FUNCTION_BLOCK "FB_Arg_Seq_1"   // FB2, GRAPH_PLUS
{ S7_Optimized_Access := 'TRUE' }
VERSION : 0.1
   VAR_INPUT
      OFF_SQ : Bool := false;   // Turn sequence off
      INIT_SQ : Bool := false;   // Set sequence to initial state
      ACK_EF : Bool := false;   // Acknowledge all errors and faults
      S_PREV : Bool := false;   // Output previous step in parameter S_NO
      S_NEXT : Bool := false;   // Indicate next step in parameter S_NO
      SW_AUTO : Bool := false;   // Automatic mode
      SW_TAP : Bool := false;   // Semiautomatic/switch with transition
      SW_TOP : Bool := false;   // Semiautomatic/ignore transition
      SW_MAN : Bool := false;   // Manual mode
      S_SEL : Int := 0;   // Select step to be output to S_NO
      S_ON : Bool := false;   // Activate step indicated in S_NO
      S_OFF : Bool := false;   // Deactivate step indicated S_NO
      T_PUSH : Bool := false;   // Enable transition to switch in semi automatic mode
      Start : Bool;
      stepTimes : Array[2..10] of Time;
      Model_Numb : Int := 3;
   END_VAR
   VAR_OUTPUT
      S_NO : Int := 0;   // Step number
      S_MORE : Bool := false;   // More steps are available and can be shown in S_NO
      S_ACTIVE : Bool := false;   // Step indicated in S_NO is active
      ERR_FLT : Bool := false;   // Interlock or supervision group error
      AUTO_ON : Bool := false;   // Automatic mode is active
      TAP_ON : Bool := false;   // Semiautomatic mode/step with transition enabled
      TOP_ON : Bool := false;   // Semiautomatic mode/ignore transition enabled
      MAN_ON : Bool := false;   // Manual mode is active
   END_VAR
   VAR
      HMI_INFO : Array[0..8] of UInt;
      IF_PAR : G7_IfParPlus_V6;
      RT_DATA : G7_RTDataPlus_V6;   // Internal data area
      Trans1 : G7_TransitionPlus_V6;   // Transition structure
      Trans2 : G7_TransitionPlus_V6;   // Transition structure
      Trans3 : G7_TransitionPlus_V6;   // Transition structure
      Trans4 : G7_TransitionPlus_V6;   // Transition structure
      Trans5 : G7_TransitionPlus_V6;   // Transition structure
      Trans6 : G7_TransitionPlus_V6;   // Transition structure
      Trans7 : G7_TransitionPlus_V6;   // Transition structure
      Trans8 : G7_TransitionPlus_V6;   // Transition structure
      Trans9 : G7_TransitionPlus_V6;   // Transition structure
      Trans10 : G7_TransitionPlus_V6;   // Transition structure
      Trans11 : G7_TransitionPlus_V6;   // Transition structure
      Trans12 : G7_TransitionPlus_V6;   // Transition structure
      Trans13 : G7_TransitionPlus_V6;   // Transition structure
      Trans14 : G7_TransitionPlus_V6;   // Transition structure
      Trans15 : G7_TransitionPlus_V6;   // Transition structure
      Trans16 : G7_TransitionPlus_V6;   // Transition structure
      Trans17 : G7_TransitionPlus_V6;   // Transition structure
      Trans18 : G7_TransitionPlus_V6;   // Transition structure
      Trans19 : G7_TransitionPlus_V6;   // Transition structure
      Trans21 : G7_TransitionPlus_V6;   // Transition structure
      "Step1: Init (Idle)" : G7_StepPlus_V6;   // Step structure
      Step2 : G7_StepPlus_V6;   // Step structure
      Step3 : G7_StepPlus_V6;   // Step structure
      Step4 : G7_StepPlus_V6;   // Step structure
      Step5 : G7_StepPlus_V6;   // Step structure
      Step6 : G7_StepPlus_V6;   // Step structure
      Step7 : G7_StepPlus_V6;   // Step structure
      Step8 : G7_StepPlus_V6;   // Step structure
      Step9 : G7_StepPlus_V6;   // Step structure
      Step10 : G7_StepPlus_V6;   // Step structure
      Step11 : G7_StepPlus_V6;   // Step structure
      Step12 : G7_StepPlus_V6;   // Step structure
      Step13 : G7_StepPlus_V6;   // Step structure
      Step14 : G7_StepPlus_V6;   // Step structure
      Step15 : G7_StepPlus_V6;   // Step structure
      Step16 : G7_StepPlus_V6;   // Step structure
      Step17 : G7_StepPlus_V6;   // Step structure
      Step18 : G7_StepPlus_V6;   // Step structure
      Step19 : G7_StepPlus_V6;   // Step structure
      SINI : Array[0..1] of USInt;
      LSTT : Array[0..19] of USInt;
      ATAJ : Array[0..19] of USInt;
      ATAB : Array[0..19] of USInt;
      PSTT : Array[0..19] of USInt;
      NSTT : Array[0..19] of USInt;
      ASSJ : Array[0..18] of USInt;
      ASSB : Array[0..18] of USInt;
      PTTS : Array[0..18] of USInt;
      NTTS : Array[0..18] of USInt;
      SW_SQTS : Array[0..18] of USInt;
      SWITCH : Array[0..1] of USInt;
      TVX : Array[0..3] of USInt;
      TTX : Array[0..3] of USInt;
      TSX : Array[0..1] of USInt;
      S00X : Array[0..1] of USInt;
      SOFFX : Array[0..1] of USInt;
      SONX : Array[0..1] of USInt;
      SAX : Array[0..1] of USInt;
      SERRX : Array[0..19] of USInt;
      SMX : Array[0..19] of USInt;
      S0X : Array[0..19] of USInt;
      S1X : Array[0..19] of USInt;
      IL_ALARM_INST : Diag_Alarm;
      SUP_ALARM_INST : Diag_Alarm;
      STEP_TIME_ALARM_INST : Diag_Alarm;
      IEC_TIMER_INST : IEC_TIMER;
      TRANSACTION_FLAG : Bool := false;
   END_VAR
   // SINI[0] := 2;
   // LSTT[0] := 255;
   // LSTT[1] := 255;
   // LSTT[2] := 255;
   // ATAJ[1] := 1;
   // ATAJ[2] := 2;
   // ATAJ[3] := 3;
   // ATAB[1] := 1;
   // ATAB[2] := 2;
   // ATAB[3] := 3;
   // PSTT[1] := 1;
   // PSTT[2] := 2;
   // PSTT[3] := 3;
   // NSTT[0] := 1;
   // NSTT[1] := 2;
   // NSTT[2] := 3;
   // ASSJ[1] := 1;
   // ASSJ[2] := 2;
   // ASSJ[3] := 3;
   // ASSB[1] := 1;
   // ASSB[2] := 2;
   // ASSB[3] := 3;
   // PTTS[0] := 255;
   // PTTS[2] := 1;
   // PTTS[3] := 2;
   // NTTS[1] := 1;
   // NTTS[2] := 2;
   // NTTS[3] := 3;
   // TVX[0] := 16#1;
   // TTX[0] := 16#1;
   // TSX[0] := 16#1;
   // S00X[0] := 16#1;
   // SOFFX[0] := 16#1;
   // SONX[0] := 16#1;
   // SAX[0] := 16#1;
   // SERRX[0] := 16#1;
   // SMX[0] := 16#1;
   // S0X[0] := 16#1;
   // S1X[0] := 16#1;
   // LSTT[3] := 255;
   // LSTT[4] := 255;
   // LSTT[5] := 255;
   // LSTT[6] := 255;
   // LSTT[7] := 255;
   // LSTT[8] := 255;
   // ATAJ[4] := 4;
   // ATAJ[5] := 5;
   // ATAJ[6] := 6;
   // ATAJ[7] := 7;
   // ATAJ[8] := 8;
   // ATAJ[9] := 9;
   // ATAB[4] := 4;
   // ATAB[5] := 5;
   // ATAB[6] := 6;
   // ATAB[7] := 7;
   // ATAB[8] := 8;
   // ATAB[9] := 9;
   // PSTT[4] := 4;
   // PSTT[5] := 5;
   // PSTT[6] := 6;
   // PSTT[7] := 7;
   // PSTT[8] := 8;
   // PSTT[9] := 9;
   // NSTT[3] := 4;
   // NSTT[4] := 5;
   // NSTT[5] := 6;
   // NSTT[6] := 7;
   // NSTT[7] := 8;
   // NSTT[8] := 9;
   // ASSJ[4] := 4;
   // ASSJ[5] := 5;
   // ASSJ[6] := 6;
   // ASSJ[7] := 7;
   // ASSJ[8] := 8;
   // ASSJ[9] := 9;
   // ASSB[4] := 4;
   // ASSB[5] := 5;
   // ASSB[6] := 6;
   // ASSB[7] := 7;
   // ASSB[8] := 8;
   // ASSB[9] := 9;
   // PTTS[4] := 3;
   // PTTS[5] := 4;
   // PTTS[6] := 5;
   // PTTS[7] := 6;
   // PTTS[8] := 7;
   // PTTS[9] := 8;
   // NTTS[4] := 4;
   // NTTS[5] := 5;
   // NTTS[6] := 6;
   // NTTS[7] := 7;
   // NTTS[8] := 8;
   // NTTS[9] := 9;
   // LSTT[10] := 255;
   // LSTT[11] := 255;
   // LSTT[12] := 255;
   // LSTT[13] := 255;
   // LSTT[14] := 255;
   // LSTT[15] := 255;
   // LSTT[16] := 255;
   // LSTT[17] := 255;
   // LSTT[18] := 255;
   // ATAJ[10] := 10;
   // ATAJ[11] := 11;
   // ATAJ[12] := 12;
   // ATAJ[13] := 13;
   // ATAJ[14] := 14;
   // ATAJ[15] := 15;
   // ATAJ[16] := 16;
   // ATAJ[17] := 17;
   // ATAJ[18] := 18;
   // ATAJ[19] := 19;
   // ATAB[0] := 10;
   // ATAB[11] := 11;
   // ATAB[12] := 12;
   // ATAB[13] := 13;
   // ATAB[14] := 14;
   // ATAB[15] := 15;
   // ATAB[16] := 16;
   // ATAB[17] := 17;
   // ATAB[18] := 18;
   // ATAB[19] := 19;
   // PSTT[11] := 10;
   // PSTT[12] := 11;
   // PSTT[13] := 12;
   // PSTT[14] := 13;
   // PSTT[15] := 14;
   // PSTT[16] := 15;
   // PSTT[17] := 16;
   // PSTT[18] := 17;
   // PSTT[19] := 18;
   // NSTT[10] := 10;
   // NSTT[11] := 11;
   // NSTT[12] := 12;
   // NSTT[13] := 13;
   // NSTT[14] := 14;
   // NSTT[15] := 15;
   // NSTT[16] := 16;
   // NSTT[17] := 17;
   // NSTT[18] := 18;
   // ASSJ[10] := 10;
   // ASSJ[11] := 11;
   // ASSJ[12] := 12;
   // ASSJ[13] := 13;
   // ASSJ[14] := 14;
   // ASSJ[15] := 15;
   // ASSJ[16] := 16;
   // ASSJ[17] := 17;
   // ASSJ[18] := 18;
   // ASSB[10] := 10;
   // ASSB[11] := 11;
   // ASSB[12] := 12;
   // ASSB[13] := 13;
   // ASSB[14] := 14;
   // ASSB[15] := 15;
   // ASSB[16] := 16;
   // ASSB[17] := 17;
   // ASSB[18] := 18;
   // PTTS[10] := 10;
   // PTTS[11] := 11;
   // PTTS[12] := 12;
   // PTTS[13] := 13;
   // PTTS[14] := 14;
   // PTTS[15] := 15;
   // PTTS[16] := 16;
   // PTTS[17] := 17;
   // PTTS[18] := 18;
   // NTTS[10] := 11;
   // NTTS[11] := 12;
   // NTTS[12] := 13;
   // NTTS[13] := 14;
   // NTTS[14] := 15;
   // NTTS[15] := 16;
   // NTTS[16] := 17;
   // NTTS[17] := 18;
   // NTTS[18] := 19;
   // SW_SQTS[1] := 1;
   // SW_SQTS[2] := 1;
   // SW_SQTS[3] := 1;
   // SW_SQTS[4] := 1;
   // SW_SQTS[5] := 1;
   // SW_SQTS[6] := 1;
   // SW_SQTS[7] := 1;
   // SW_SQTS[8] := 1;
   // SW_SQTS[9] := 1;
   // SW_SQTS[10] := 2;
   // SW_SQTS[11] := 2;
   // SW_SQTS[12] := 2;
   // SW_SQTS[13] := 2;
   // SW_SQTS[14] := 2;
   // SW_SQTS[15] := 2;
   // SW_SQTS[16] := 2;
   // SW_SQTS[17] := 2;
   // SW_SQTS[18] := 2;
BEGIN
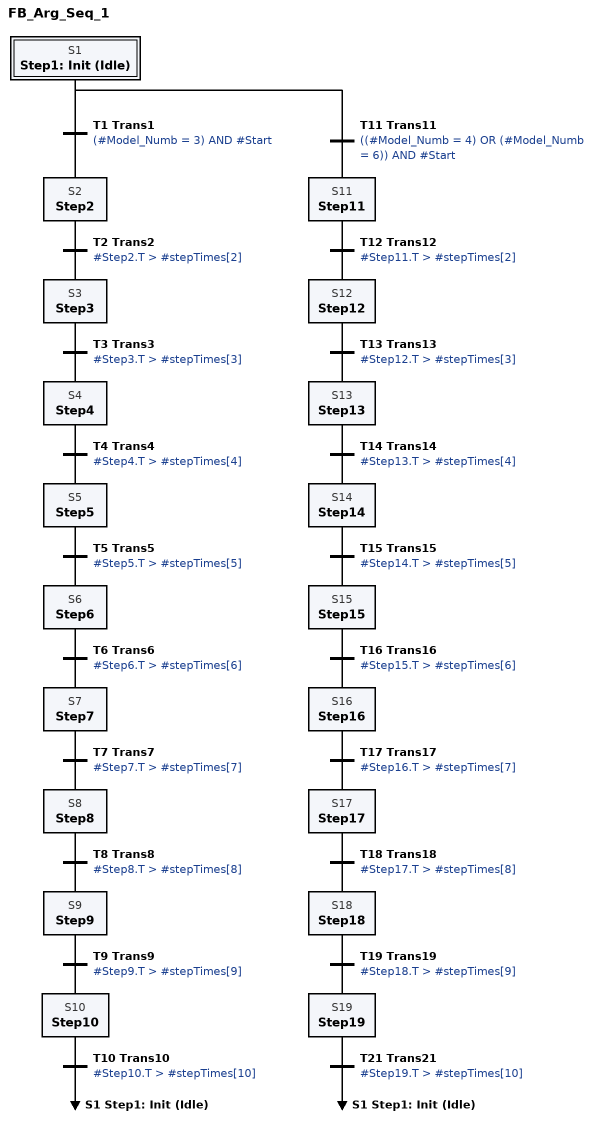
   // sequencer 1
   INITIAL_STEP "Step1: Init (Idle)":   // S1, max time T#10S, warning time T#7S
   END_STEP
   TRANSITION Trans1 FROM "Step1: Init (Idle)" TO Step2   // T1
      := (#Model_Numb = 3) AND #Start;
   END_TRANSITION
   TRANSITION Trans11 FROM "Step1: Init (Idle)" TO Step11   // T11
      := ((#Model_Numb = 4) OR (#Model_Numb = 6)) AND #Start;
   END_TRANSITION
   STEP Step2:   // S2, max time T#10S, warning time T#7S
   END_STEP
   TRANSITION Trans2 FROM Step2 TO Step3   // T2
      := #Step2.T > #stepTimes[2];
   END_TRANSITION
   STEP Step3:   // S3, max time T#10S, warning time T#7S
   END_STEP
   TRANSITION Trans3 FROM Step3 TO Step4   // T3
      := #Step3.T > #stepTimes[3];
   END_TRANSITION
   STEP Step4:   // S4, max time T#10S, warning time T#7S
   END_STEP
   TRANSITION Trans4 FROM Step4 TO Step5   // T4
      := #Step4.T > #stepTimes[4];
   END_TRANSITION
   STEP Step5:   // S5, max time T#10S, warning time T#7S
   END_STEP
   TRANSITION Trans5 FROM Step5 TO Step6   // T5
      := #Step5.T > #stepTimes[5];
   END_TRANSITION
   STEP Step6:   // S6, max time T#10S, warning time T#7S
   END_STEP
   TRANSITION Trans6 FROM Step6 TO Step7   // T6
      := #Step6.T > #stepTimes[6];
   END_TRANSITION
   STEP Step7:   // S7, max time T#10S, warning time T#7S
   END_STEP
   TRANSITION Trans7 FROM Step7 TO Step8   // T7
      := #Step7.T > #stepTimes[7];
   END_TRANSITION
   STEP Step8:   // S8, max time T#10S, warning time T#7S
   END_STEP
   TRANSITION Trans8 FROM Step8 TO Step9   // T8
      := #Step8.T > #stepTimes[8];
   END_TRANSITION
   STEP Step9:   // S9, max time T#10S, warning time T#7S
   END_STEP
   TRANSITION Trans9 FROM Step9 TO Step10   // T9
      := #Step9.T > #stepTimes[9];
   END_TRANSITION
   STEP Step10:   // S10, max time T#10S, warning time T#7S
   END_STEP
   TRANSITION Trans10 FROM Step10 TO "Step1: Init (Idle)"   // T10, jump
      := #Step10.T > #stepTimes[10];
   END_TRANSITION
   STEP Step11:   // S11, max time T#10S, warning time T#7S
   END_STEP
   TRANSITION Trans12 FROM Step11 TO Step12   // T12
      := #Step11.T > #stepTimes[2];
   END_TRANSITION
   STEP Step12:   // S12, max time T#10S, warning time T#7S
   END_STEP
   TRANSITION Trans13 FROM Step12 TO Step13   // T13
      := #Step12.T > #stepTimes[3];
   END_TRANSITION
   STEP Step13:   // S13, max time T#10S, warning time T#7S
   END_STEP
   TRANSITION Trans14 FROM Step13 TO Step14   // T14
      := #Step13.T > #stepTimes[4];
   END_TRANSITION
   STEP Step14:   // S14, max time T#10S, warning time T#7S
   END_STEP
   TRANSITION Trans15 FROM Step14 TO Step15   // T15
      := #Step14.T > #stepTimes[5];
   END_TRANSITION
   STEP Step15:   // S15, max time T#10S, warning time T#7S
   END_STEP
   TRANSITION Trans16 FROM Step15 TO Step16   // T16
      := #Step15.T > #stepTimes[6];
   END_TRANSITION
   STEP Step16:   // S16, max time T#10S, warning time T#7S
   END_STEP
   TRANSITION Trans17 FROM Step16 TO Step17   // T17
      := #Step16.T > #stepTimes[7];
   END_TRANSITION
   STEP Step17:   // S17, max time T#10S, warning time T#7S
   END_STEP
   TRANSITION Trans18 FROM Step17 TO Step18   // T18
      := #Step17.T > #stepTimes[8];
   END_TRANSITION
   STEP Step18:   // S18, max time T#10S, warning time T#7S
   END_STEP
   TRANSITION Trans19 FROM Step18 TO Step19   // T19
      := #Step18.T > #stepTimes[9];
   END_TRANSITION
   STEP Step19:   // S19, max time T#10S, warning time T#7S
   END_STEP
   TRANSITION Trans21 FROM Step19 TO "Step1: Init (Idle)"   // T21, jump
      := #Step19.T > #stepTimes[10];
   END_TRANSITION
END_FUNCTION_BLOCK

FUNCTION "FC_ARG_1" : Void   // FC1, FBD
{ S7_Optimized_Access := 'TRUE' }
VERSION : 0.1
   VAR_OUTPUT
      Ready_new_car : Bool;
   END_VAR
   VAR_TEMP
      stepTimes : Array[2..10] of Time;
      i : Int;
      Random_Time : Time;   // Random Time between 0sec to 10sec
      Start : Bool;
      Stop : Bool;
      status1_RandFunc : Word;
      status2_RandFunc : Word;
      temp : Byte;
      error_RandFunc : Bool;
   END_VAR
   VAR CONSTANT
      sequenceNO : Int := 9;
   END_VAR
BEGIN

REGION Network 1 (SCL): Man Mode Data Handling
   IF "DB_Process_Var".Man_Mode = TRUE THEN
       "DB_Process_Var".Car_Type_Selected := "DB_HMI".dropdown_selection;
   END_IF;
END_REGION

REGION Network 2 (SCL): Auto Mode Data Handling
   IF "DB_Process_Var".Auto_Mode = TRUE THEN
       "DB_HMI".dropdown_selection := 0;
       "DB_Process_Var".Car_Type_Selected := "DB_PLC5_Receiving".ReceivingBoxForward.Type;
   END_IF;
   IF "DB_HMI".ARG1_Seq1_Cmd_Auto OR "DB_HMI".Global_Cmd_Auto THEN
       "DB_HMI".dropdown_selection := 0;
       "DB_Process_Var".Car_Type_Selected := 0;
   END_IF;
END_REGION

REGION Network 3 (SCL): Load Time Date based on Car Type
       CASE "DB_Process_Var".Car_Type_Selected OF
           3:
               "DB_Profile"."time" := "DB_Profile".time_Red;
           4:
               "DB_Profile"."time" := "DB_Profile".time_Green;
           6:
               "DB_Profile"."time" := "DB_Profile".time_Blue;
       END_CASE;
END_REGION

REGION Network 4 (SCL): Switch from selected to inProduction
   IF "IDB_Arg_Seq_1_DB".Trans1.TS = TRUE OR "IDB_Arg_Seq_1_DB".Trans11.TS = TRUE THEN
       IF "DB_Process_Var".Car_Type_Selected = 3 THEN
           "DB_Process_Var".Car_Type_inProduction := 3;
           "DB_Process_Var".Car_Type_inProduction_Text := 'Red';
           "DB_HMI".ARG1_Seq1_inProduction := 3;
       ELSIF "DB_Process_Var".Car_Type_Selected = 4 THEN
           "DB_Process_Var".Car_Type_inProduction := 4;
           "DB_Process_Var".Car_Type_inProduction_Text := 'Green';
           "DB_HMI".ARG1_Seq1_inProduction := 4;
       ELSIF "DB_Process_Var".Car_Type_Selected = 6 THEN
           "DB_Process_Var".Car_Type_inProduction := 6;
           "DB_Process_Var".Car_Type_inProduction_Text := 'Blue';
           "DB_HMI".ARG1_Seq1_inProduction := 6;
       END_IF;
   END_IF;
END_REGION

REGION Network 5 (SCL): Create Random Time Values for the selected Steps
   IF "IDB_Arg_Seq_1_DB".Trans1.TS = TRUE OR "IDB_Arg_Seq_1_DB".Trans11.TS = TRUE THEN
       FOR #i := 2 TO 10 DO
           //Red
           IF "DB_HMI".ARG1_Seq1_DelaySelect_Red[#i] = TRUE THEN;
               "DB_Sim".Delta_T_Red[#i] := "LGF_RandomRange_Dint"(minValue := 0, maxValue := 10000, error => #error_RandFunc, status => #status1_RandFunc, subfunctionStatus => #status2_RandFunc);
           ELSE
               "DB_Sim".Delta_T_Red[#i] := T#0s;
           END_IF;
           //Green
           IF "DB_HMI".ARG1_Seq1_DelaySelect_Green[#i] = TRUE THEN
               "DB_Sim".Delta_T_Green[#i] := "LGF_RandomRange_Dint"(minValue := 0, maxValue := 10000, error => #error_RandFunc, status => #status1_RandFunc, subfunctionStatus => #status2_RandFunc);
           ELSE
               "DB_Sim".Delta_T_Green[#i] := T#0s;
           END_IF;
           //Blue
           IF "DB_HMI".ARG1_Seq1_DelaySelect_Blue[#i] = TRUE THEN
               "DB_Sim".Delta_T_Blue[#i] := "LGF_RandomRange_Dint"(minValue := 0, maxValue := 10000, error => #error_RandFunc, status => #status1_RandFunc, subfunctionStatus => #status2_RandFunc);
           ELSE
               "DB_Sim".Delta_T_Blue[#i] := T#0s;
           END_IF;
       END_FOR;
   END_IF;

   IF "DB_HMI".ARG1_Seq1_Cmd_DelayReset = TRUE THEN
       FOR #i := 2 TO 10 DO
           "DB_HMI".ARG1_Seq1_DelaySelect_Red[#i] := false;
           "DB_HMI".ARG1_Seq1_DelaySelect_Green[#i] := false;
           "DB_HMI".ARG1_Seq1_DelaySelect_Blue[#i] := false;
       END_FOR;
   END_IF;
END_REGION

REGION Network 6 (SCL): Add Delay Time to Step Time
   FOR #i := 2 TO 10 DO
       IF "DB_HMI".dropdown_selection = 3 OR "DB_PLC5_Receiving".ReceivingBoxForward.Type = 3 THEN
           "DB_Process_Var".Step_Times[#i] := T_ADD(IN1 := "DB_Profile"."time"[#i], IN2 := "DB_Sim".Delta_T_Red[#i]);
       ELSIF "DB_HMI".dropdown_selection = 4 OR "DB_PLC5_Receiving".ReceivingBoxForward.Type = 4 THEN
           "DB_Process_Var".Step_Times[#i] := T_ADD(IN1 := "DB_Profile"."time"[#i], IN2 := "DB_Sim".Delta_T_Green[#i]);
       ELSIF "DB_HMI".dropdown_selection = 6 OR "DB_PLC5_Receiving".ReceivingBoxForward.Type = 6 THEN
           "DB_Process_Var".Step_Times[#i] := T_ADD(IN1 := "DB_Profile"."time"[#i], IN2 := "DB_Sim".Delta_T_Blue[#i]);
       END_IF;
   END_FOR;
END_REGION

REGION Network 7: Auto Mode select
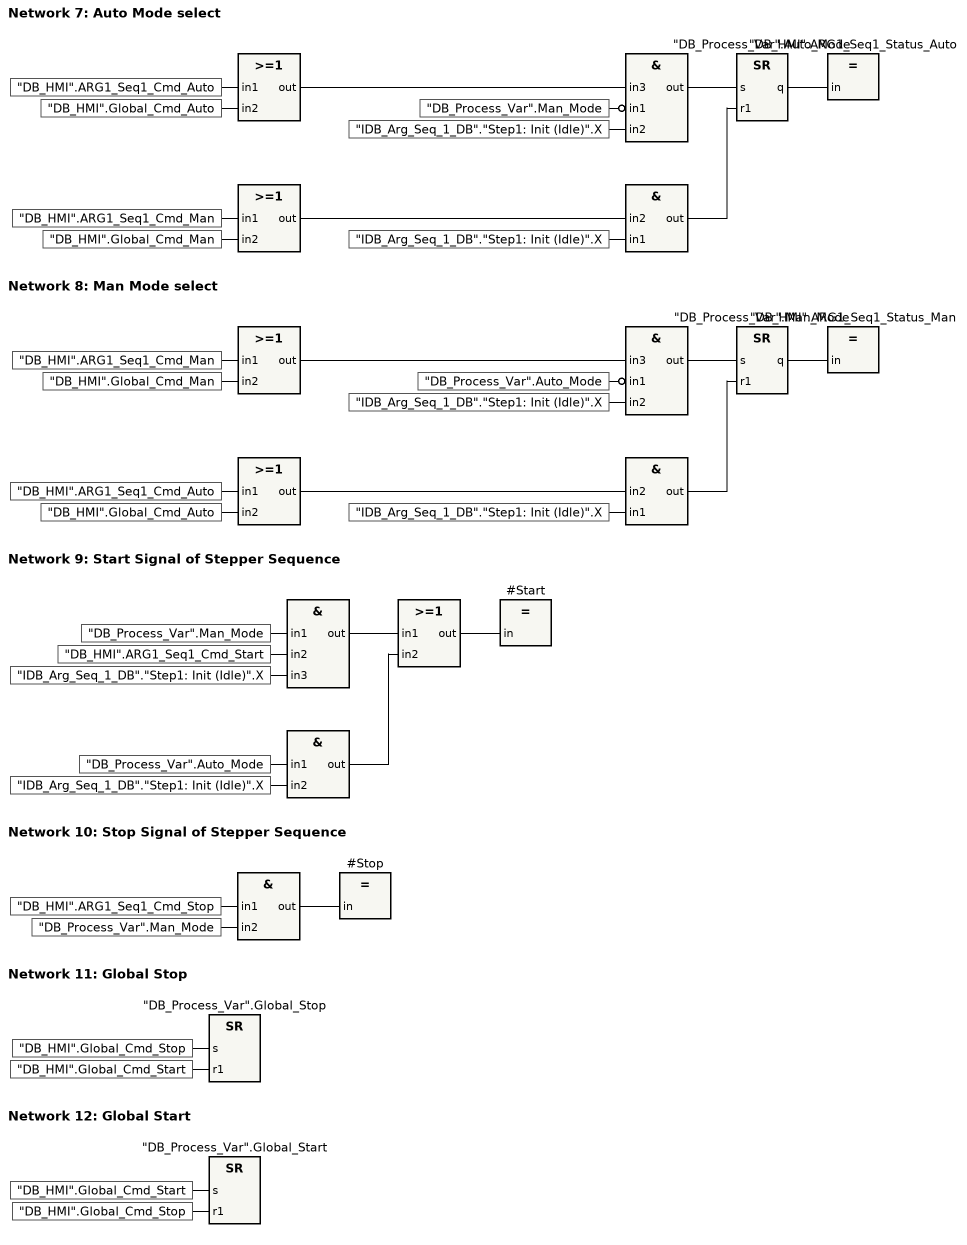
   IF ("DB_HMI".ARG1_Seq1_Cmd_Auto OR "DB_HMI".Global_Cmd_Auto) AND NOT "DB_Process_Var".Man_Mode AND "IDB_Arg_Seq_1_DB"."Step1: Init (Idle)".X THEN
       "DB_Process_Var".Auto_Mode := TRUE;   // SR flip-flop
   END_IF;
   IF ("DB_HMI".ARG1_Seq1_Cmd_Man OR "DB_HMI".Global_Cmd_Man) AND "IDB_Arg_Seq_1_DB"."Step1: Init (Idle)".X THEN
       "DB_Process_Var".Auto_Mode := FALSE;
   END_IF;
   "DB_HMI".ARG1_Seq1_Status_Auto := "DB_Process_Var".Auto_Mode;
END_REGION

REGION Network 8: Man Mode select
   IF ("DB_HMI".ARG1_Seq1_Cmd_Man OR "DB_HMI".Global_Cmd_Man) AND NOT "DB_Process_Var".Auto_Mode AND "IDB_Arg_Seq_1_DB"."Step1: Init (Idle)".X THEN
       "DB_Process_Var".Man_Mode := TRUE;   // SR flip-flop
   END_IF;
   IF ("DB_HMI".ARG1_Seq1_Cmd_Auto OR "DB_HMI".Global_Cmd_Auto) AND "IDB_Arg_Seq_1_DB"."Step1: Init (Idle)".X THEN
       "DB_Process_Var".Man_Mode := FALSE;
   END_IF;
   "DB_HMI".ARG1_Seq1_Status_Man := "DB_Process_Var".Man_Mode;
END_REGION

REGION Network 9: Start Signal of Stepper Sequence
   #Start := ("DB_Process_Var".Man_Mode AND "DB_HMI".ARG1_Seq1_Cmd_Start AND "IDB_Arg_Seq_1_DB"."Step1: Init (Idle)".X) OR ("DB_Process_Var".Auto_Mode AND "IDB_Arg_Seq_1_DB"."Step1: Init (Idle)".X);
END_REGION

REGION Network 10: Stop Signal of Stepper Sequence
   #Stop := "DB_HMI".ARG1_Seq1_Cmd_Stop AND "DB_Process_Var".Man_Mode;
END_REGION

REGION Network 11: Global Stop
   IF "DB_HMI".Global_Cmd_Stop THEN
       "DB_Process_Var".Global_Stop := TRUE;   // SR flip-flop
   END_IF;
   IF "DB_HMI".Global_Cmd_Start THEN "DB_Process_Var".Global_Stop := FALSE; END_IF;
END_REGION

REGION Network 12: Global Start
   IF "DB_HMI".Global_Cmd_Start THEN
       "DB_Process_Var".Global_Start := TRUE;   // SR flip-flop
   END_IF;
   IF "DB_HMI".Global_Cmd_Stop THEN "DB_Process_Var".Global_Start := FALSE; END_IF;
END_REGION

REGION Network 13 (SCL): Reset Type Selection
   IF "DB_HMI".ARG1_Seq1_Cmd_Stop = TRUE THEN
       "DB_PLC5_Receiving".ReceivingBoxForward.Type := 0;
       "DB_HMI".ARG1_Seq1_inProduction := 0;
       "DB_Process_Var".ReadyNewCar := TRUE;
   END_IF;
END_REGION

REGION Network 14: Call FB with Stepper Sequence
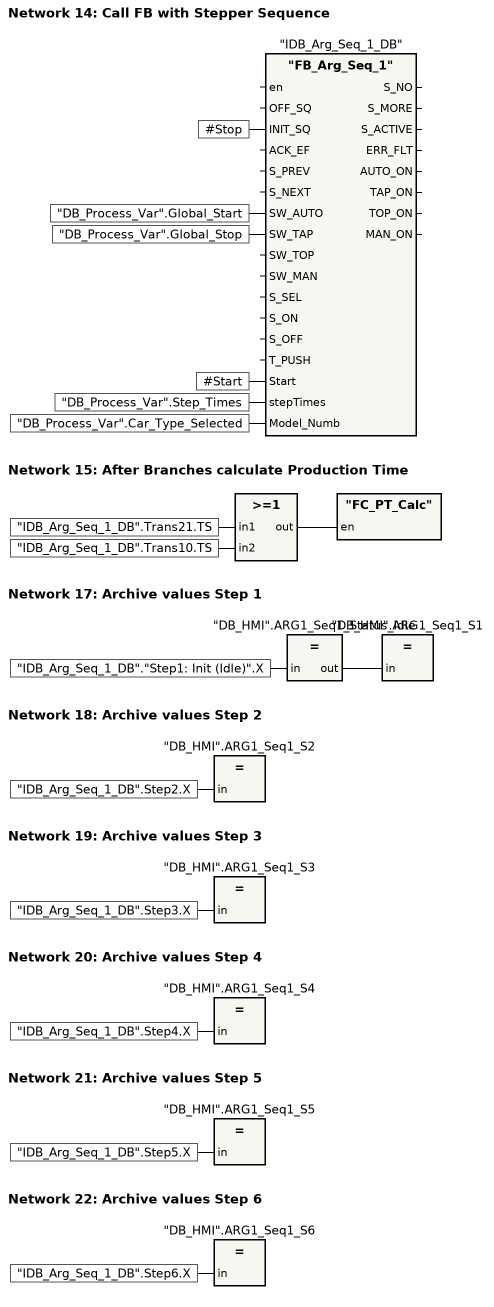
   "IDB_Arg_Seq_1_DB"(INIT_SQ := #Stop,   // "FB_Arg_Seq_1"
                      SW_AUTO := "DB_Process_Var".Global_Start,
                      SW_TAP := "DB_Process_Var".Global_Stop,
                      Start := #Start,
                      stepTimes := "DB_Process_Var".Step_Times,
                      Model_Numb := "DB_Process_Var".Car_Type_Selected);
END_REGION

REGION Network 15: After Branches calculate Production Time
   IF "IDB_Arg_Seq_1_DB".Trans21.TS OR "IDB_Arg_Seq_1_DB".Trans10.TS THEN "FC_PT_Calc"(); END_IF;
END_REGION

REGION Network 16 (SCL): Send Idle to previous Station
   IF "IDB_Arg_Seq_1_DB"."Step1: Init (Idle)".X = TRUE THEN
       "DB_PLC5_Sending".SendBox.Station_Idle := TRUE;
   ELSE
       "DB_PLC5_Sending".SendBox.Station_Idle := FALSE;
   END_IF;
END_REGION

REGION Network 17: Archive values Step 1
   "DB_HMI".ARG1_Seq1_Status_Idle := "IDB_Arg_Seq_1_DB"."Step1: Init (Idle)".X;
   "DB_HMI".ARG1_Seq1_S1 := "IDB_Arg_Seq_1_DB"."Step1: Init (Idle)".X;
END_REGION

REGION Network 18: Archive values Step 2
   "DB_HMI".ARG1_Seq1_S2 := "IDB_Arg_Seq_1_DB".Step2.X;
END_REGION

REGION Network 19: Archive values Step 3
   "DB_HMI".ARG1_Seq1_S3 := "IDB_Arg_Seq_1_DB".Step3.X;
END_REGION

REGION Network 20: Archive values Step 4
   "DB_HMI".ARG1_Seq1_S4 := "IDB_Arg_Seq_1_DB".Step4.X;
END_REGION

REGION Network 21: Archive values Step 5
   "DB_HMI".ARG1_Seq1_S5 := "IDB_Arg_Seq_1_DB".Step5.X;
END_REGION

REGION Network 22: Archive values Step 6
   "DB_HMI".ARG1_Seq1_S6 := "IDB_Arg_Seq_1_DB".Step6.X;
END_REGION

REGION Network 23: Archive values Step 7
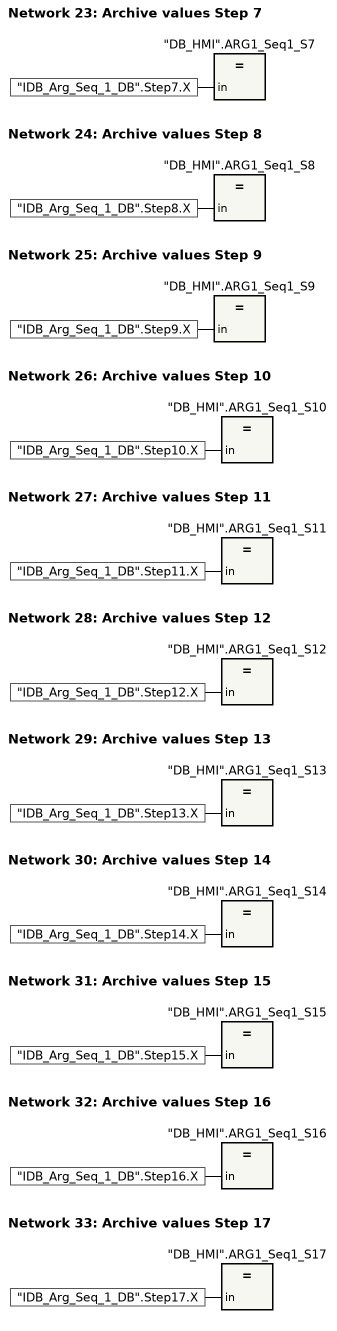
   "DB_HMI".ARG1_Seq1_S7 := "IDB_Arg_Seq_1_DB".Step7.X;
END_REGION

REGION Network 24: Archive values Step 8
   "DB_HMI".ARG1_Seq1_S8 := "IDB_Arg_Seq_1_DB".Step8.X;
END_REGION

REGION Network 25: Archive values Step 9
   "DB_HMI".ARG1_Seq1_S9 := "IDB_Arg_Seq_1_DB".Step9.X;
END_REGION

REGION Network 26: Archive values Step 10
   "DB_HMI".ARG1_Seq1_S10 := "IDB_Arg_Seq_1_DB".Step10.X;
END_REGION

REGION Network 27: Archive values Step 11
   "DB_HMI".ARG1_Seq1_S11 := "IDB_Arg_Seq_1_DB".Step11.X;
END_REGION

REGION Network 28: Archive values Step 12
   "DB_HMI".ARG1_Seq1_S12 := "IDB_Arg_Seq_1_DB".Step12.X;
END_REGION

REGION Network 29: Archive values Step 13
   "DB_HMI".ARG1_Seq1_S13 := "IDB_Arg_Seq_1_DB".Step13.X;
END_REGION

REGION Network 30: Archive values Step 14
   "DB_HMI".ARG1_Seq1_S14 := "IDB_Arg_Seq_1_DB".Step14.X;
END_REGION

REGION Network 31: Archive values Step 15
   "DB_HMI".ARG1_Seq1_S15 := "IDB_Arg_Seq_1_DB".Step15.X;
END_REGION

REGION Network 32: Archive values Step 16
   "DB_HMI".ARG1_Seq1_S16 := "IDB_Arg_Seq_1_DB".Step16.X;
END_REGION

REGION Network 33: Archive values Step 17
   "DB_HMI".ARG1_Seq1_S17 := "IDB_Arg_Seq_1_DB".Step17.X;
END_REGION

REGION Network 34: Archive values Step 18
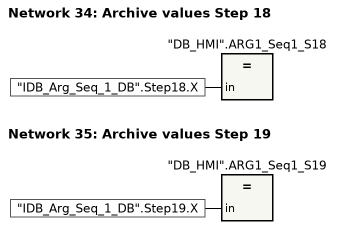
   "DB_HMI".ARG1_Seq1_S18 := "IDB_Arg_Seq_1_DB".Step18.X;
END_REGION

REGION Network 35: Archive values Step 19
   "DB_HMI".ARG1_Seq1_S19 := "IDB_Arg_Seq_1_DB".Step19.X;
END_REGION

REGION Network 36 (SCL): Set Busy
   IF
       "IDB_Arg_Seq_1_DB".Step2.X OR
       "IDB_Arg_Seq_1_DB".Step3.X OR
       "IDB_Arg_Seq_1_DB".Step4.X OR
       "IDB_Arg_Seq_1_DB".Step5.X OR
       "IDB_Arg_Seq_1_DB".Step6.X OR
       "IDB_Arg_Seq_1_DB".Step7.X OR
       "IDB_Arg_Seq_1_DB".Step8.X OR
       "IDB_Arg_Seq_1_DB".Step9.X OR
       "IDB_Arg_Seq_1_DB".Step10.X OR
       "IDB_Arg_Seq_1_DB".Step11.X OR
       "IDB_Arg_Seq_1_DB".Step12.X OR
       "IDB_Arg_Seq_1_DB".Step13.X OR
       "IDB_Arg_Seq_1_DB".Step14.X OR
       "IDB_Arg_Seq_1_DB".Step15.X OR
       "IDB_Arg_Seq_1_DB".Step16.X OR
       "IDB_Arg_Seq_1_DB".Step17.X OR
       "IDB_Arg_Seq_1_DB".Step18.X OR
       "IDB_Arg_Seq_1_DB".Step19.X THEN
       "DB_HMI".ARG1_Seq1_Status_Busy := TRUE;
   ELSIF "IDB_Arg_Seq_1_DB"."Step1: Init (Idle)".X THEN
       "DB_HMI".ARG1_Seq1_Status_Busy := FALSE;
   END_IF;
END_REGION

REGION Network 37 (SCL): When Stepper Sequence runs completely
   IF "IDB_Arg_Seq_1_DB".Trans10.TS = TRUE OR "IDB_Arg_Seq_1_DB".Trans21.TS = TRUE THEN
       "DB_Process_Var".Branch_Complete := TRUE;
       "DB_Process_Var".Car_Type_Ready := "DB_Process_Var".Car_Type_inProduction;
       "DB_Process_Var".Car_Type_inProduction := 0;
       "DB_Process_Var".Car_Type_inProduction_Text := '';
       "DB_Process_Var".Car_ReadyToShift := TRUE;
       "DB_HMI".ARG1_Seq1_inProduction := 0;
   END_IF;
   IF "IDB_Arg_Seq_1_DB".Trans1.TS = TRUE OR "IDB_Arg_Seq_1_DB".Trans11.TS = TRUE THEN
       "DB_Process_Var".Branch_Complete := FALSE;
       "DB_Process_Var".ReadyNewCar := 0;
   END_IF;
END_REGION

REGION Network 38 (SCL): Write Data in the Sending Box
   //IF "DB_Process_Var".Branch_Complete = TRUE AND "DB_PLC5_Receiving".ReceivingBox.Station_Idle = TRUE THEN
   IF "IDB_Arg_Seq_1_DB".Trans10.TS = TRUE OR "IDB_Arg_Seq_1_DB".Trans21.TS = TRUE THEN
       "DB_PLC5_Sending".SendBoxForward.Planned_PT_Red := "DB_HMI".ARG1_Seq1_Calculated_PT_Red;
       "DB_PLC5_Sending".SendBoxForward.Planned_PT_Green := "DB_HMI".ARG1_Seq1_Calculated_PT_Green;
       "DB_PLC5_Sending".SendBoxForward.Planned_PT_Blue := "DB_HMI".ARG1_Seq1_Calculated_PT_Blue;

       "DB_PLC5_Sending".SendBoxForward.Measuered_PT_Red := "DB_HMI".ARG1_Seq1_Messured_PT_Red;
       "DB_PLC5_Sending".SendBoxForward.Measuered_PT_Green := "DB_HMI".ARG1_Seq1_Messured_PT_Green;
       "DB_PLC5_Sending".SendBoxForward.Measuered_PT_Blue := "DB_HMI".ARG1_Seq1_Messured_PT_Blue;

       "DB_PLC5_Sending".SendBoxForward.Type := "DB_Process_Var".Car_Type_Ready;

       "DB_PLC5_Receiving".ReceivingBoxForward.Type := 0;

       "DB_HMI".ARG1_Seq1_inProduction := 0;
   END_IF;
END_REGION

REGION Network 39 (SCL): Reset Receiving Car Typ
   //IF "IDB_Arg_Seq_1_DB".Trans1.TS = TRUE OR "IDB_Arg_Seq_1_DB".Trans11.TS THEN
       //"DB_PLC5_Receiving".ReceivingBoxForward.Type := 0;
   //END_IF;
END_REGION

REGION Network 40 (SCL): When car is shifted
   IF "DB_Process_Var".Data_Put_Done = TRUE THEN
       "DB_Process_Var".Car_Type_Ready := 0;
       "DB_PLC5_Sending".SendBoxForward.Type := 0;
       "DB_Process_Var".Car_ReadyToShift := FALSE;
       "DB_HMI".ARG1_Seq1_inProduction := 0;
       "DB_Process_Var".ReadyNewCar := 1;
       //"DB_PLC5_Receiving".ReceivingBoxForward.Type := 0;
   END_IF;
END_REGION
END_FUNCTION

FUNCTION "FC_Com" : Void   // FC2, FBD
{ S7_Optimized_Access := 'TRUE' }
VERSION : 0.1
BEGIN

REGION Network 1: Communication PLC1 -> PLC2
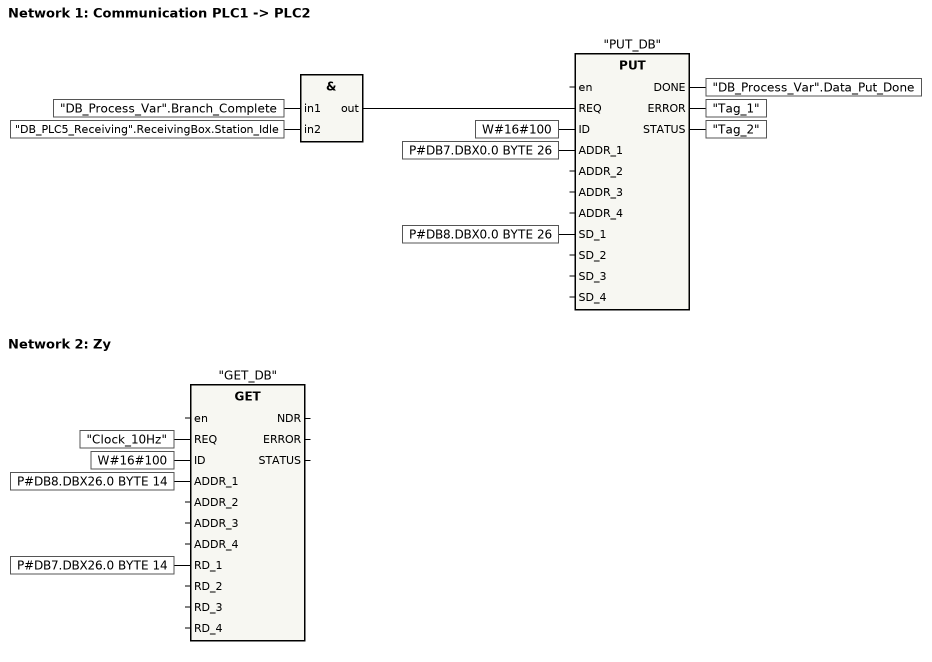
   "PUT_DB"(REQ := "DB_Process_Var".Branch_Complete AND "DB_PLC5_Receiving".ReceivingBox.Station_Idle,   // PUT
            ID := W#16#100,
            ADDR_1 := P#DB7.DBX0.0 BYTE 26,
            SD_1 := P#DB8.DBX0.0 BYTE 26,
            DONE => "DB_Process_Var".Data_Put_Done,
            ERROR => "Tag_1",
            STATUS => "Tag_2");
END_REGION

REGION Network 2: Zy
   "GET_DB"(REQ := "Clock_10Hz", ID := W#16#100, ADDR_1 := P#DB8.DBX26.0 BYTE 14, RD_1 := P#DB7.DBX26.0 BYTE 14);   // GET
END_REGION
END_FUNCTION

FUNCTION "FC_PT_Calc" : Void   // FC3, SCL
{ S7_Optimized_Access := 'TRUE' }
VERSION : 0.1
   VAR_TEMP
      i : Int;
   END_VAR
   VAR CONSTANT
      sequenceNO : Int := 9;
      Null : Time := T#0MS;
   END_VAR
BEGIN
   "DB_HMI".ARG1_Seq1_Calculated_PT_Red := #Null;
   "DB_HMI".ARG1_Seq1_Calculated_PT_Green := #Null;
   "DB_HMI".ARG1_Seq1_Calculated_PT_Blue := #Null;

   "DB_HMI".ARG1_Seq1_Messured_PT_Red := #Null;
   "DB_HMI".ARG1_Seq1_Messured_PT_Green := #Null;
   "DB_HMI".ARG1_Seq1_Messured_PT_Blue := #Null;